DATA_BLOCK "DB_Z201_HMI"   // DB2010
{ S7_Optimized_Access := 'FALSE' }
VERSION : 0.1
   VAR
      tAlm : Struct   // HMI Alarms
         tE : Struct   // Emergency alarms
            xMainEmergency : Bool := TRUE;   // A122KE1.Main emergency ON {X|X|X|X|O}
            xSpare_1 : Bool := TRUE;
            xSpare_2 : Bool := TRUE;
            xSpare_3 : Bool := TRUE;
            xSpare_4 : Bool := TRUE;
            xSpare_5 : Bool := TRUE;
            xLocalMain1 : Bool := TRUE;   // A118SB1.Emergency localization MCC1201 {X|X|X|X|O}
            xLocalMain2 : Bool := TRUE;   // A118SB2.Emergency localization CS4201 {X|X|X|X|O}
            xLocalMain3 : Bool := TRUE;   // M204SSB3.Emergency localization M204S {X|X|X|X|O}
            xLocalMain4 : Bool := TRUE;   // M204SSB4.Emergency localization M204S {X|X|X|X|O}
            xLocalMain5 : Bool := FALSE;   // M211SB1.Emergency localization M211 {X|X|X|X|O}
            xLocalMain6 : Bool := FALSE;   // M211SB2.Emergency localization M211 {X|X|X|X|O}
            xLocalMain7 : Bool := FALSE;   // M218SB1.Emergency localization M218 {X|X|X|X|O}
            xLocalMain8 : Bool := FALSE;   // M218SB2.Emergency localization M218 {X|X|X|X|O}
            xLocalMain9 : Bool := FALSE;   // M214SB1.Emergency localization M214 {X|X|X|X|O}
            xLocalMain10 : Bool := FALSE;   // M214SB2.Emergency localization M214 {X|X|X|X|O}
            xLocalMain11 : Bool := FALSE;   // M203SB1.Emergency localization M203 {X|X|X|X|O}
            xLocalMain12 : Bool := FALSE;   // AxxSBx.Emergency localization Spare {X|X|X|X|O}
            xLocalMain13 : Bool := FALSE;   // AxxSBx.Emergency localization Spare {X|X|X|X|O}
            xSpare_19 : Bool := FALSE;
            xEmergencyONArea201 : Bool := FALSE;   // Emergency ON Area 201
            xEmergencyONArea301 : Bool := FALSE;   // Emergency ON Area 301
            xEmergencyONArea302 : Bool := FALSE;   // Emergency ON Area 302
            xEmergencyONArea501 : Bool := FALSE;   // Emergency ON Area 501
            xEmergencyONArea601 : Bool := FALSE;   // Emergency ON Area 601
            xEmergencyONArea701 : Bool := FALSE;   // Emergency ON Area 701
            xEmergencyONArea303 : Bool := FALSE;   // Emergency ON Area 303
            xSpare_27 : Bool := FALSE;
            xSpare_28 : Bool := FALSE;
            xSpare_29 : Bool := FALSE;
            xSpare_30 : Bool := FALSE;
            xSpare_31 : Bool := FALSE;
         END_STRUCT;
         tS : Struct   // Stopping faults
            xZ300NotReady : Bool := FALSE;   // Area 300 is not ready {X|X|X|X|O}
            xSpare_1 : Bool := FALSE;
            xSpare_2 : Bool := FALSE;
            xSpare_3 : Bool := FALSE;
            xSpare_4 : Bool := FALSE;
            xSpare_5 : Bool := FALSE;
            xSpare_6 : Bool := FALSE;
            xSpare_7 : Bool := FALSE;
            xSpare_8 : Bool := FALSE;
            xSpare_9 : Bool := FALSE;
            xSpare_10 : Bool := FALSE;
            xSpare_11 : Bool := FALSE;
            xSpare_12 : Bool := FALSE;
            xSpare_13 : Bool := FALSE;
            xSpare_14 : Bool := FALSE;
            xSpare_15 : Bool := FALSE;
            xSpare_16 : Bool := FALSE;
            xSpare_17 : Bool := FALSE;
            xSpare_18 : Bool := FALSE;
            xSpare_19 : Bool := FALSE;
            xSpare_20 : Bool := FALSE;
            xSpare_21 : Bool := FALSE;
            xSpare_22 : Bool := FALSE;
            xSpare_23 : Bool := FALSE;
            xSpare_24 : Bool := FALSE;
            xSpare_25 : Bool := FALSE;
            xSpare_26 : Bool := FALSE;
            xSpare_27 : Bool := FALSE;
            xSpare_28 : Bool := FALSE;
            xSpare_29 : Bool := FALSE;
            xSpare_30 : Bool := FALSE;
            xSpare_31 : Bool := FALSE;
         END_STRUCT;
         tF : Struct   // Faults
            xPowerFailure230vAux : Bool := FALSE;   // NU_A10QF1/2.Power failure 230v auxiliary / R13QF1.R13QF2.Power failure 230v auxiliary
            xPowerSupply24vLogic : Bool := FALSE;   // A109QF2.Power supply 24v logic / R18QF3.Power supply 24v logic
            xPowerSupply24vLogic2 : Bool := FALSE;   // A109QF3.Power supply 24v logic / R18QF4.Power supply 24v logic
            xPowerSuppluyOut24vUnderUpsEmOk : Bool := FALSE;   // A108QF5.Out24vUnderUpsEmOk / R18AP1.Redundancy 24v ok
            xPowerSupply24vLogic3 : Bool := FALSE;   // NU_A19QF1.Power supply 24v logic
            xPowerSupply24vLogic4 : Bool := FALSE;   // NU_A19QF2.Power supply 24v logic
            xPowerSuppluyOut24vUnderEmOk : Bool := FALSE;   // A108QF6.Out24vUnderEmOk
            xSpare_7 : Bool := FALSE;
            xPowerSupply24vDrive2 : Bool := FALSE;   // NU_A20QF4.Power Supply 24V Drive
            xSpare_9 : Bool := FALSE;
            xDriveSupply2 : Bool := FALSE;   // A137QM1.Drive Supply
            xSpare_11 : Bool := FALSE;
            xM216FanProtection : Bool;   // M216.A141QM1.Fan protection
            xM216FanFeedback : Bool;   // M216.A141KM1.Feedback rotation / M250.R12KM1.Feedback rotation
            xM209FanFeedback : Bool;   // M209.A178KM1.Feedback Rotation
            xSpare_15 : Bool;
            xSpare_16 : Bool;
            xSpare_17 : Bool;   // R204SP1.Compressed air presence cutting bridges
            xSpare_18 : Bool;
            xSpare_19 : Bool;
            xSpare_20 : Bool := FALSE;
            xSpare_21 : Bool := FALSE;
            xSpare_22 : Bool := FALSE;
            xSpare_23 : Bool := FALSE;
            xSpare_24 : Bool := FALSE;
            xSpare_25 : Bool := FALSE;
            xSpare_26 : Bool := FALSE;
            xSpare_27 : Bool := FALSE;
            xSpare_28 : Bool := FALSE;
            xSpare_29 : Bool := FALSE;
            xSpare_30 : Bool := FALSE;
            xSpare_31 : Bool := FALSE;
         END_STRUCT;
         tW : Struct   // Warnings
            xSpare_0 : Bool := FALSE;
            xSpare_1 : Bool := FALSE;
            xSpare_2 : Bool := FALSE;
            xSpare_3 : Bool := FALSE;
            xSpare_4 : Bool := FALSE;
            xSpare_5 : Bool := FALSE;
            xSpare_6 : Bool := FALSE;
            xSpare_7 : Bool := FALSE;
            xSpare_8 : Bool := FALSE;
            xSpare_9 : Bool := FALSE;
            xSpare_10 : Bool := FALSE;
            xSpare_11 : Bool := FALSE;
            xSpare_12 : Bool := FALSE;
            xSpare_13 : Bool := FALSE;
            xSpare_14 : Bool := FALSE;
            xSpare_15 : Bool := FALSE;
            xSpare_16 : Bool := FALSE;
            xSpare_17 : Bool := FALSE;
            xSpare_18 : Bool := FALSE;
            xSpare_19 : Bool := FALSE;
            xSpare_20 : Bool := FALSE;
            xSpare_21 : Bool := FALSE;
            xSpare_22 : Bool := FALSE;
            xSpare_23 : Bool := FALSE;
            xSpare_24 : Bool := FALSE;
            xSpare_25 : Bool := FALSE;
            xSpare_26 : Bool := FALSE;
            xSpare_27 : Bool := FALSE;
            xSpare_28 : Bool := FALSE;
            xSpare_29 : Bool := FALSE;
            xSpare_30 : Bool := FALSE;
            xSpare_31 : Bool := FALSE;
         END_STRUCT;
      END_STRUCT;
      tHMR : Struct   // HMI Read
         xSpare0 : Bool;
         xSpare1 : Bool;
         xSpare2 : Bool;
         xSpare3 : Bool;
         xSpare4 : Bool;
         xSpare5 : Bool;
         xSpare6 : Bool;
         xSpare7 : Bool;
         xSpare8 : Bool;
         xSpare9 : Bool;
         xSpare10 : Bool;
         xSpare11 : Bool;
         xSpare12 : Bool;
         xSpare13 : Bool;
         xSpare14 : Bool;
         xZoneAlarm : Bool := FALSE;   // Zone alarm {X|X|X|X|O}
         xSpare16 : Bool;
         xSpare17 : Bool;
         xSpare18 : Bool;
         xSpare19 : Bool;
         xSpare20 : Bool;
         xSpare21 : Bool;
         xSpare22 : Bool;
         xSpare23 : Bool;
         xSpare24 : Bool;
         xSpare25 : Bool;
         xSpare26 : Bool;
         xSpare27 : Bool;
         xSpare28 : Bool;
         xSpare29 : Bool;
         xSpare30 : Bool;
         xSpare31 : Bool;
         xSpare : Array[0..15] of Bool;
         iSpare0 : Int;
         iSpare1 : Int;
         iSpare2 : Int;
         iSpare3 : Int;
         iSpare4 : Int;
         iSpare5 : Int;
         iSpare6 : Int;
         iSpare7 : Int;
         iSpare8 : Int;
         iSpare9 : Int;
         iSpare10 : Int;
         iSpare11 : Int;
         iSpare12 : Int;
         iSpare13 : Int;
         iSpare14 : Int;
         iSpare15 : Int;
         iSpare16 : Int;
         dSpare0 : DInt;
         dZoneState : DInt := 1024;   // Zone status (1=CycleON 2=StopCyc 4=CycleReq 8=StopReq 1024=E-Stop) {X|X|X|X|O} / HMI Alarms
         dCabinetStatusMCC : DInt := 1;   // Cabinet status MCC1201 (1=OK;2=General power alarm;3=Local power alarm) {X|X|X|X|O} / HMI Write
         dDistanceFromSnaproll_cmm_M209 : DInt;   // Distance from snaproll [mm/100] {mm/100|mm|0|60000|M}
         dDistanceFromSnaproll_cmm_M216 : DInt;   // Distance from snaproll [mm/100] {mm/100|mm|0|60000|M}
         dSpare5 : DInt;
         dSpare6 : DInt;
         dSpare7 : DInt;
         dSpare8 : DInt;
         dSpare9 : DInt;
         dSpare10 : DInt;
         dSpare11 : DInt;
         dSpare12 : DInt;
         dSpare13 : DInt;
         dSpare14 : DInt;
         dSpare15 : DInt;
         rSpare0 : Real;
         rSpare1 : Real;
         rSpare2 : Real;
         rSpare3 : Real;
         rSpare4 : Real;
         rSpare5 : Real;
         rSpare6 : Real;
         rSpare7 : Real;
         rSpare8 : Real;
         tManCmd : Struct
            xFdbkRunFw : Bool;   // Feedback rotation FW all conveyors {x|x|x|x|O}
            xSpare1 : Bool;
            xSpare2 : Bool;
            xSpare3 : Bool;
            xSpare4 : Bool;
            xSpare5 : Bool;
            xSpare6 : Bool;
            xSpare7 : Bool;
            xSpare8 : Bool;
            xSpare9 : Bool;
            xSpare10 : Bool;
            xSpare11 : Bool;
            xSpare12 : Bool;
            xSpare13 : Bool;
            xSpare14 : Bool;
            xSpare15 : Bool;
            xSpare : Array[0..15] of Bool;
         END_STRUCT;
      END_STRUCT;
      tHMW : Struct   // HMI Write
         xSpare0 : Bool;
         xSpare1 : Bool;
         xSpare2 : Bool;
         xSpare3 : Bool;
         xSpare4 : Bool;
         xStartCycleRequest : Bool := FALSE;   // Start cycle request {X|X|X|X|O}
         xStopCycleRequest : Bool := FALSE;   // Stop cycle request {X|X|X|X|O}
         xForceStopCycle : Bool := FALSE;   // Force stop cycle {X|X|X|X|O}
         xSpare8 : Bool;
         xEnabledChipsBlowerM216 : Bool;   // Chips Blower M216 Enabled {X|X|X|X|O}
         xEnabledChipsBlowerM209 : Bool;   // Chips Blower M209 Enabled {X|X|X|X|O}
         xUpdateDistSnap_M209 : Bool;   // Update distance from snap roll {x|x|x|x|M}
         xUpdateDistSnap_M216 : Bool;
         xSpare13 : Bool;
         xEnableManualCommand : Bool;   // Enable Disable Manual command {x|x|x|x|O}
         xFaultsReset : Bool := FALSE;   // Reset faults {X|X|X|X|O}
         xGeneralReset : Bool := FALSE;   // General reset {X|X|X|X|M}
         xSpare17 : Bool;
         xSpare18 : Bool;
         xSpare19 : Bool;
         xSpare20 : Bool;
         xSpare21 : Bool;
         xSpare22 : Bool;
         xSpare23 : Bool;
         xSpare24 : Bool;
         xSpare25 : Bool;
         xSpare26 : Bool;
         xSpare27 : Bool;
         xSpare28 : Bool;
         xSpare29 : Bool;
         xSpare30 : Bool;
         xSpare31 : Bool;
         xSpare : Array[0..15] of Bool;
         iSpare0 : Int;
         iSpare1 : Int;
         iSpare2 : Int;
         iSpare3 : Int;
         iSpare4 : Int;
         iSpare5 : Int;
         iSpare6 : Int;
         iSpare7 : Int;
         iSpare8 : Int;
         iSpare9 : Int;
         iSpare10 : Int;
         iSpare11 : Int;
         iSpare12 : Int;
         iSpare13 : Int;
         iSpare14 : Int;
         iSpare15 : Int;
         iSpare16 : Int;
         dDistanceFromSnaproll_cmm_M209 : DInt;   // Distance from snaproll [mm/100] [mm/100] {mm/100|mm|0|60000|M}
         dDistanceFromSnaproll_cmm_M216 : DInt;   // Distance from snaproll [mm/100] [mm/100] {mm/100|mm|0|60000|M}
         dSpare2 : DInt;
         dSpare3 : DInt;
         dSpare4 : DInt;
         dSpare5 : DInt;
         dSpare6 : DInt;
         dSpare7 : DInt;
         dSpare8 : DInt;
         dSpare9 : DInt;
         dSpare10 : DInt;
         dSpare11 : DInt;
         dSpare12 : DInt;
         dSpare13 : DInt;
         dSpare14 : DInt;
         dSpare15 : DInt;
         dSpare16 : DInt;
         rSpare0 : Real;
         rSpare1 : Real;
         rSpare2 : Real;
         rSpare3 : Real;
         rSpare4 : Real;
         rSpare5 : Real;
         rSpare6 : Real;
         rSpare7 : Real;
         rSpare8 : Real;
         tManCmd : Struct
            xRunFw : Bool;   // Rotation FW all conveyors {x|x|x|x|O}
            xSpare1 : Bool;
            xSpare2 : Bool;
            xSpare3 : Bool;
            xSpare4 : Bool;
            xSpare5 : Bool;
            xSpare6 : Bool;
            xSpare7 : Bool;
            xSpare8 : Bool;
            xSpare9 : Bool;
            xSpare10 : Bool;
            xSpare11 : Bool;
            xSpare12 : Bool;
            xSpare13 : Bool;
            xSpare14 : Bool;
            xSpare15 : Bool;
            xSpare16 : Bool;
            xSpare17 : Bool;
            xSpare18 : Bool;
            xSpare19 : Bool;
            xSpare20 : Bool;
            xSpare21 : Bool;
            xSpare22 : Bool;
            xSpare23 : Bool;
            xSpare24 : Bool;
            xSpare25 : Bool;
            xSpare26 : Bool;
            xSpare27 : Bool;
            xSpare28 : Bool;
            xSpare29 : Bool;
            xSpare30 : Bool;
            xSpare31 : Bool;
         END_STRUCT;
      END_STRUCT;
   END_VAR
BEGIN
END_DATA_BLOCK

DATA_BLOCK "DB_ZUPS_HMI"   // DB2012
{ S7_Optimized_Access := 'FALSE' }
VERSION : 0.1
   VAR
      tAlm : Struct   // HMI Alarms
         tE : Struct   // Emergency alarms
            xSpare_0 : Bool := TRUE;
            xMainEmergencyUPS : Bool := TRUE;   // A117KE1.Main emergency UPS ON {X|X|X|X|O}
            xLocalUPS1 : Bool := TRUE;   // AxxSB1.Emergency localization MCC1201 {X|X|X|X|O}
            xLocalUPS2 : Bool := TRUE;   // M204S_SB1.Emergency localization M204S {X|X|X|X|O}
            xLocalUPS3 : Bool := TRUE;   // M204S_SB2.Emergency localization M204S {X|X|X|X|O}
            xLocalUPS4 : Bool := TRUE;   // CS4201A117SB1.Emergency localization spare {X|X|X|X|O}
            xLocalUpS5 : Bool := TRUE;   // AxxSBx.Emergency localization spare {X|X|X|X|O}
            xSpare_7 : Bool := TRUE;
            xSpare_8 : Bool := TRUE;
            xSpare_9 : Bool := TRUE;
            xSpare_10 : Bool := FALSE;
            xSpare_11 : Bool := FALSE;
            xSpare_12 : Bool := FALSE;
            xSpare_13 : Bool := FALSE;
            xSpare_14 : Bool := FALSE;
            xSpare_15 : Bool := FALSE;
            xSpare_16 : Bool := FALSE;
            xSpare_17 : Bool := FALSE;
            xSpare_18 : Bool := FALSE;
            xSpare_19 : Bool := FALSE;
            xSpare_20 : Bool := FALSE;
            xSpare_21 : Bool := FALSE;
            xSpare_22 : Bool := FALSE;
            xSpare_23 : Bool := FALSE;
            xSpare_24 : Bool := FALSE;
            xSpare_25 : Bool := FALSE;
            xSpare_26 : Bool := FALSE;
            xSpare_27 : Bool := FALSE;
            xSpare_28 : Bool := FALSE;
            xSpare_29 : Bool := FALSE;
            xSpare_30 : Bool := FALSE;
            xSpare_31 : Bool := FALSE;
         END_STRUCT;
         tS : Struct   // Stopping faults
            xSpare_0 : Bool := FALSE;
            xSpare_1 : Bool := FALSE;
            xSpare_2 : Bool := FALSE;
            xSpare_3 : Bool := FALSE;
            xSpare_4 : Bool := FALSE;
            xSpare_5 : Bool := FALSE;
            xSpare_6 : Bool := FALSE;
            xSpare_7 : Bool := FALSE;
            xSpare_8 : Bool := FALSE;
            xSpare_9 : Bool := FALSE;
            xSpare_10 : Bool := FALSE;
            xSpare_11 : Bool := FALSE;
            xSpare_12 : Bool := FALSE;
            xSpare_13 : Bool := FALSE;
            xSpare_14 : Bool := FALSE;
            xSpare_15 : Bool := FALSE;
            xSpare_16 : Bool := FALSE;
            xSpare_17 : Bool := FALSE;
            xSpare_18 : Bool := FALSE;
            xSpare_19 : Bool := FALSE;
            xSpare_20 : Bool := FALSE;
            xSpare_21 : Bool := FALSE;
            xSpare_22 : Bool := FALSE;
            xSpare_23 : Bool := FALSE;
            xSpare_24 : Bool := FALSE;
            xSpare_25 : Bool := FALSE;
            xSpare_26 : Bool := FALSE;
            xSpare_27 : Bool := FALSE;
            xSpare_28 : Bool := FALSE;
            xSpare_29 : Bool := FALSE;
            xSpare_30 : Bool := FALSE;
            xSpare_31 : Bool := FALSE;
         END_STRUCT;
         tF : Struct   // Faults
            xSpare_0 : Bool := FALSE;   // R13QF1.R13QF2.Power failure 230v auxiliary
            xSpare_1 : Bool := FALSE;   // R18QF3.Power supply 24v logic
            xSpare_2 : Bool := FALSE;   // R18QF4.Power supply 24v logic
            xSpare_3 : Bool := FALSE;   // R18AP1.Redundancy 24v ok
            xSpare_4 : Bool := FALSE;
            xSpare_5 : Bool := FALSE;
            xSpare_6 : Bool := FALSE;
            xPowerSupply24vDrive1 : Bool := FALSE;   // A110QF2.Power Supply 24V Drive
            xSpare_8 : Bool := FALSE;
            xDriveSupply1 : Bool := FALSE;   // A136QM1.Drive Supply
            xSpare_10 : Bool := FALSE;
            xSpare_11 : Bool := FALSE;
            xSpare_12 : Bool;
            xSpare_13 : Bool;   // M250.R12KM1.Feedback rotation
            xSpare_14 : Bool;
            xSpare_15 : Bool;
            xSpare_16 : Bool;
            xSpare_17 : Bool;   // R204SP1.Compressed air presence cutting bridges
            xSpare_18 : Bool;
            xSpare_19 : Bool;
            xSpare_20 : Bool := FALSE;
            xSpare_21 : Bool := FALSE;
            xSpare_22 : Bool := FALSE;
            xSpare_23 : Bool := FALSE;
            xSpare_24 : Bool := FALSE;
            xSpare_25 : Bool := FALSE;
            xSpare_26 : Bool := FALSE;
            xSpare_27 : Bool := FALSE;
            xSpare_28 : Bool := FALSE;
            xSpare_29 : Bool := FALSE;
            xSpare_30 : Bool := FALSE;
            xSpare_31 : Bool := FALSE;
         END_STRUCT;
         tW : Struct   // Warnings
            xSpare_0 : Bool := FALSE;
            xSpare_1 : Bool := FALSE;
            xSpare_2 : Bool := FALSE;
            xSpare_3 : Bool := FALSE;
            xSpare_4 : Bool := FALSE;
            xSpare_5 : Bool := FALSE;
            xSpare_6 : Bool := FALSE;
            xSpare_7 : Bool := FALSE;
            xSpare_8 : Bool := FALSE;
            xSpare_9 : Bool := FALSE;
            xSpare_10 : Bool := FALSE;
            xSpare_11 : Bool := FALSE;
            xSpare_12 : Bool := FALSE;
            xSpare_13 : Bool := FALSE;
            xSpare_14 : Bool := FALSE;
            xSpare_15 : Bool := FALSE;
            xSpare_16 : Bool := FALSE;
            xSpare_17 : Bool := FALSE;
            xSpare_18 : Bool := FALSE;
            xSpare_19 : Bool := FALSE;
            xSpare_20 : Bool := FALSE;
            xSpare_21 : Bool := FALSE;
            xSpare_22 : Bool := FALSE;
            xSpare_23 : Bool := FALSE;
            xSpare_24 : Bool := FALSE;
            xSpare_25 : Bool := FALSE;
            xSpare_26 : Bool := FALSE;
            xSpare_27 : Bool := FALSE;
            xSpare_28 : Bool := FALSE;
            xSpare_29 : Bool := FALSE;
            xSpare_30 : Bool := FALSE;
            xSpare_31 : Bool := FALSE;
         END_STRUCT;
      END_STRUCT;
      tHMR : Struct   // HMI Read
         xSpare0 : Bool;
         xSpare1 : Bool;
         xSpare2 : Bool;
         xSpare3 : Bool;
         xSpare4 : Bool;
         xSpare5 : Bool;
         xSpare6 : Bool;
         xSpare7 : Bool;
         xSpare8 : Bool;
         xSpare9 : Bool;
         xSpare10 : Bool;
         xSpare11 : Bool;
         xSpare12 : Bool;
         xSpare13 : Bool;
         xSpare14 : Bool;
         xZoneAlarm : Bool := FALSE;   // Zone alarm {X|X|X|X|O}
         xSpare16 : Bool;
         xSpare17 : Bool;
         xSpare18 : Bool;
         xSpare19 : Bool;
         xSpare20 : Bool;
         xSpare21 : Bool;
         xSpare22 : Bool;
         xSpare23 : Bool;
         xSpare24 : Bool;
         xSpare25 : Bool;
         xSpare26 : Bool;
         xSpare27 : Bool;
         xSpare28 : Bool;
         xSpare29 : Bool;
         xSpare30 : Bool;
         xSpare31 : Bool;
         xSpare : Array[0..15] of Bool;
         iSpare0 : Int;
         iSpare1 : Int;
         iSpare2 : Int;
         iSpare3 : Int;
         iSpare4 : Int;
         iSpare5 : Int;
         iSpare6 : Int;
         iSpare7 : Int;
         iSpare8 : Int;
         iSpare9 : Int;
         iSpare10 : Int;
         iSpare11 : Int;
         iSpare12 : Int;
         iSpare13 : Int;
         iSpare14 : Int;
         iSpare15 : Int;
         iSpare16 : Int;
         dSpare0 : DInt;
         dZoneState : DInt := 1024;   // Zone status (1=CycleON 2=StopCyc 4=CycleReq 8=StopReq 1024=E-Stop) {X|X|X|X|O} / HMI Alarms
         dSpare2 : DInt;
         dSpare3 : DInt;
         dSpare4 : DInt;
         dSpare5 : DInt;
         dSpare6 : DInt;
         dSpare7 : DInt;
         dSpare8 : DInt;
         dSpare9 : DInt;
         dSpare10 : DInt;
         dSpare11 : DInt;
         dSpare12 : DInt;
         dSpare13 : DInt;
         dSpare14 : DInt;
         dSpare15 : DInt;
         rSpare0 : Real;
         rSpare1 : Real;
         rSpare2 : Real;
         rSpare3 : Real;
         rSpare4 : Real;
         rSpare5 : Real;
         rSpare6 : Real;
         rSpare7 : Real;
         rSpare8 : Real;
         tManCmd : Struct
            xSpare0 : Bool;
            xSpare1 : Bool;
            xSpare2 : Bool;
            xSpare3 : Bool;
            xSpare4 : Bool;
            xSpare5 : Bool;
            xSpare6 : Bool;
            xSpare7 : Bool;
            xSpare8 : Bool;
            xSpare9 : Bool;
            xSpare10 : Bool;
            xSpare11 : Bool;
            xSpare12 : Bool;
            xSpare13 : Bool;
            xSpare14 : Bool;
            xSpare15 : Bool;
            xSpare : Array[0..15] of Bool;
         END_STRUCT;
      END_STRUCT;
      tHMW : Struct   // HMI Write
         xSpare0 : Bool;
         xSpare1 : Bool;
         xSpare2 : Bool;
         xSpare3 : Bool;
         xSpare4 : Bool;
         xStartCycleRequest : Bool := FALSE;   // Start cycle request {X|X|X|X|O}
         xStopCycleRequest : Bool := FALSE;   // Stop cycle request {X|X|X|X|O}
         xForceStopCycle : Bool := FALSE;   // Force stop cycle {X|X|X|X|O}
         xSpare8 : Bool;
         xSpare9 : Bool;
         xSpare10 : Bool;
         xSpare11 : Bool;
         xSpare12 : Bool;
         xSpare13 : Bool;
         xSpare14 : Bool;
         xFaultsReset : Bool := FALSE;   // Reset faults {X|X|X|X|O}
         xSpare16 : Bool := FALSE;
         xSpare17 : Bool;
         xSpare18 : Bool;
         xSpare19 : Bool;
         xSpare20 : Bool;
         xSpare21 : Bool;
         xSpare22 : Bool;
         xSpare23 : Bool;
         xSpare24 : Bool;
         xSpare25 : Bool;
         xSpare26 : Bool;
         xSpare27 : Bool;
         xSpare28 : Bool;
         xSpare29 : Bool;
         xSpare30 : Bool;
         xSpare31 : Bool;
         xSpare : Array[0..15] of Bool;
         iSpare0 : Int;
         iSpare1 : Int;
         iSpare2 : Int;
         iSpare3 : Int;
         iSpare4 : Int;
         iSpare5 : Int;
         iSpare6 : Int;
         iSpare7 : Int;
         iSpare8 : Int;
         iSpare9 : Int;
         iSpare10 : Int;
         iSpare11 : Int;
         iSpare12 : Int;
         iSpare13 : Int;
         iSpare14 : Int;
         iSpare15 : Int;
         iSpare16 : Int;
         dSpare0 : DInt;
         dSpare1 : DInt;
         dSpare2 : DInt;
         dSpare3 : DInt;
         dSpare4 : DInt;
         dSpare5 : DInt;
         dSpare6 : DInt;
         dSpare7 : DInt;
         dSpare8 : DInt;
         dSpare9 : DInt;
         dSpare10 : DInt;
         dSpare11 : DInt;
         dSpare12 : DInt;
         dSpare13 : DInt;
         dSpare14 : DInt;
         dSpare15 : DInt;
         dSpare16 : DInt;
         rSpare0 : Real;
         rSpare1 : Real;
         rSpare2 : Real;
         rSpare3 : Real;
         rSpare4 : Real;
         rSpare5 : Real;
         rSpare6 : Real;
         rSpare7 : Real;
         rSpare8 : Real;
         tManCmd : Struct
            xSpare0 : Bool;
            xSpare1 : Bool;
            xSpare2 : Bool;
            xSpare3 : Bool;
            xSpare4 : Bool;
            xSpare5 : Bool;
            xSpare6 : Bool;
            xSpare7 : Bool;
            xSpare8 : Bool;
            xSpare9 : Bool;
            xSpare10 : Bool;
            xSpare11 : Bool;
            xSpare12 : Bool;
            xSpare13 : Bool;
            xSpare14 : Bool;
            xSpare15 : Bool;
            xSpare16 : Bool;
            xSpare17 : Bool;
            xSpare18 : Bool;
            xSpare19 : Bool;
            xSpare20 : Bool;
            xSpare21 : Bool;
            xSpare22 : Bool;
            xSpare23 : Bool;
            xSpare24 : Bool;
            xSpare25 : Bool;
            xSpare26 : Bool;
            xSpare27 : Bool;
            xSpare28 : Bool;
            xSpare29 : Bool;
            xSpare30 : Bool;
            xSpare31 : Bool;
         END_STRUCT;
      END_STRUCT;
   END_VAR
BEGIN
END_DATA_BLOCK

// folder: TaskMedium

DATA_BLOCK "FB_OptManager_V1_00_IDB"   // DB7
{ S7_Optimized_Access := 'TRUE' }
VERSION : 0.1
// stored: InstanceOfName FB_OptManager_V1.00
"FB_OptManager_V1.00"
BEGIN
END_DATA_BLOCK

DATA_BLOCK "GP_OB_Initialize_Medium_IDB"   // DB9
{ S7_Optimized_Access := 'TRUE' }
AUTHOR : Cigliutt
FAMILY : GP
VERSION : 1.1
// stored: InstanceOfName GP_OB_Initialize
"GP_OB_Initialize"
BEGIN
END_DATA_BLOCK

DATA_BLOCK "GP_OB_Initialize_Slow_IDB"   // DB10
{ S7_Optimized_Access := 'TRUE' }
AUTHOR : Cigliutt
FAMILY : GP
VERSION : 1.1
// stored: InstanceOfName GP_OB_Initialize
"GP_OB_Initialize"
BEGIN
END_DATA_BLOCK

DATA_BLOCK "FB_Snaproll_V1_00_IDB"   // DB21
{ S7_Optimized_Access := 'TRUE' }
VERSION : 0.1
// stored: InstanceOfName FB_Snaproll_V1.00
"FB_Snaproll_V1.00"
BEGIN
END_DATA_BLOCK

DATA_BLOCK "FB_CommunicationZ300_V1.00_DB_1"   // DB25
{ S7_Optimized_Access := 'TRUE' }
VERSION : 0.1
// stored: InstanceOfName FB_CommunicationZ300_V1.00
"FB_CommunicationZ300_V1.00"
BEGIN
END_DATA_BLOCK

DATA_BLOCK "FB_CommunicationZ300_V1.00_DB"   // DB28
{ S7_Optimized_Access := 'TRUE' }
VERSION : 0.1
// stored: InstanceOfName FB_CommunicationZ300_V1.00
"FB_CommunicationZ300_V1.00"
BEGIN
END_DATA_BLOCK

DATA_BLOCK "FB_Defects_Add_Medium_V1_00_IDB"   // DB36
{ S7_Optimized_Access := 'TRUE' }
VERSION : 0.1
// stored: InstanceOfName FB_Defects_Add_V1.00
"FB_Defects_Add_V1.00"
BEGIN
END_DATA_BLOCK

// folder: TaskSlow

DATA_BLOCK "FB_Digitizer_2_V1_00_IDB"   // DB11
{ S7_Optimized_Access := 'TRUE' }
VERSION : 0.1
// stored: InstanceOfName FB_Digitizer_V1.00
"FB_Digitizer_V1.00"
BEGIN
END_DATA_BLOCK

DATA_BLOCK "FB_Digitizer_1_V1_00_IDB"   // DB12
{ S7_Optimized_Access := 'TRUE' }
VERSION : 0.1
// stored: InstanceOfName FB_Digitizer_V1.00
"FB_Digitizer_V1.00"
BEGIN
END_DATA_BLOCK

DATA_BLOCK "Z200"   // DB13
{ S7_Optimized_Access := 'TRUE' }
VERSION : 0.1
   VAR
      tmON_24Vdc : "UDT_IECTON_V1.00";   // Presence 24Vdc timer / 24VDC ok delayed timer
      ST_xZoneError : Bool := FALSE;   // Zone error / Zone is in error
      ST_xFaultsEnabled : Bool := TRUE;   // Faults enabled
      ST_xZoneFaults : Bool := TRUE;   // Cumulative of zone faults / Zone is in faults
      ST_xZoneStoppingFaults : Bool := FALSE;   // Cumulative of zone stopping faults / Zone is in stopping faults
      ST_xOutputEnabledM250Fan : Bool;   // Output enable M250 fan
      ST_xOutputEnabledM272Chips : Bool;   // Output enable M272 chips blower
      ST_xOutputEnabledM220Brush : Bool;   // Output enable M272 chips blower
      ST_xZoneWarnings : Bool := FALSE;   // Cumulative of zone warning / Zone is in warning
      ST_xCycleON : Bool := TRUE;   // Zone in cycle ON / Cycle ON
      ST_xConditionOKStopCycle : Bool := TRUE;   // Condition ok to accept stop cycle
      ST_xCycleONDelayed : Bool := TRUE;   // Cycle ON delayed
      ST_xConditionOkPhaseAdvancement : Bool := FALSE;   // Condition ok for phase advancement
      ST_xConditionOkCycleON : Bool := FALSE;   // Condition ok for cycle ON
      ST_xMachineReset : Bool := FALSE;   // Machine reset request
      ST_xPLC1 : Bool := TRUE;   // This is PLC 1
      ST_xPLC2 : Bool := FALSE;   // This is PLC 2
      ST_xThisPlcActive : Bool := TRUE;   // This PLC is active
      ST_xStartCycleRequest : Bool := FALSE;   // Request start cycle
      ST_xStopCycleRequest : Bool := FALSE;   // Request stop cycle
      ST_xM209GlassBreak : Bool;   // M272 Chips blower glass break
      ST_xM203GlassBreak : Bool;   // M272 Chips blower glass break
      OSR_xStartCycle : Bool := FALSE;   // OSR start cycle
      OSR_xStopCycle : Bool := FALSE;   // OSR stop cycle
      OSR_xForceStopCycle : Bool := FALSE;   // OSR force stop cycle
      OSR_xChipsBlowerON : Bool;   // OSR chips blower on
      OSR_xSBResetAnomaly : Bool;   // OSR reset anomaly
      OS_xStartCycle : Bool := FALSE;   // OS start cycle
      OS_xStopCycle : Bool := FALSE;   // OS stop cycle
      OS_xForceStopCycle : Bool := FALSE;   // OS force stop cycle
      OS_xChipsBlowerON : Bool;   // OS chips blower on
      OS_xCpuActive : Bool;   // OS Cpu active
      OSR_xCpuActive : Bool;   // OSR Cpu active
      ST_xStopCycleAccepted : Bool := FALSE;   // Stop cycle accepted
      AUX_tmON_M250FanFeedback : "UDT_IECTON_V1.00";   // M250 Fan feedback anomaly
      tOutputs : Struct
         xPLC1On : Bool;   // o.A195AP1.A255HL4.EnableCPUA
         xPLC2On : Bool;   // o.A195AP1.A255HL5.EnableCPUB
         xEmergencyON : Bool;   // o.A195AP1.A255HL1/1A.EmergencyON
         xSafetiesON : Bool;   // o.A195AP1.A255HL3.SafetiesON
         xHLResetAnomaly : Bool;   // o.A195AP1.A207SB1.HLResetAnomalyZ200
         xHAAlarm : Bool;   // o.A401AP1.A416HA1.Alarm
      END_STRUCT;
      tInputs : Struct
         xPowerSupply230vAux : Bool := FALSE;   // i.A195AP1.A10QF1/2.PowerFailure230VAuxiliary / i.R195AP1.R13QF1/2.PowerFailure230VAuxiliary
         xRedundancy24vOk1 : Bool;   // i.R195AP1.R18AP1.Redundacy24VOk / i.A195AP1.A18AP1.Redundancy24VOk
         xPowerSupply24vProt1 : Bool;
         xPowerSupply24vProt2 : Bool;
         xProtectionCommandsAnomalies : Bool := FALSE;   // i.A195AP1.A18QF3.PowerSupply24VLogic / i.R195AP1.R18QF3.PowerSupply24VLogic
         xProtectionCommandsInternalInput : Bool := FALSE;   // i.A195AP1.A18QF4.PowerSupply24VLogic / i.R195AP1.R18QF4.PowerSupply24VLogic
         xProtectionCommandsInternalOutput : Bool := FALSE;   // i.A195AP1.A19QF1.PowerSupply24VLogic / i.R195AP1.R18QF4.PowerSupply24VLogic
         xProtectionCommandsExternalInput : Bool := FALSE;   // i.A195AP1.A19QF2.PowerSupply24VLogic / i.R195AP1.R18QF4.PowerSupply24VLogic
         xMainEmergencyON : Bool := FALSE;   // i.A195AP1.A45KE1.MainEmergencyON / i.R195AP1.R18QF4.PowerSupply24VLogic
         xCPUAEnabled : Bool := FALSE;   // i.A151AP1.Selection CPU A / i.R150AP1.CPU A Enabled
         xCPUBEnabled : Bool := TRUE;   // i.A151AP1.Selection CPU B / i.R150AP1.CPU B Enabled
         xCPUARecognition : Bool := FALSE;   // i.A151AP1.Recognition CPU A / i.R150AP1.Recognition CPU A
         xCPUBRecognition : Bool := FALSE;   // i.A151AP1.Recognition CPU B / i.R150AP1.Recognition CPU B
         xFeedbackSwitch : Bool;
         xFeedbackAbilitationCPU_B : Bool;
         xCompressedAirPresence : Bool;
         xSBResetAnomalyZ200 : Bool;   // i.A195AP1.A207SB1.ResetAnomalyZ200
      END_STRUCT;
   END_VAR
BEGIN
END_DATA_BLOCK

DATA_BLOCK "FB_DigitizerManager_V1_00_IDB"   // DB15
{ S7_Optimized_Access := 'TRUE' }
VERSION : 0.1
// stored: InstanceOfName FB_DigitizerManager_V1.00
"FB_DigitizerManager_V1.00"
BEGIN
END_DATA_BLOCK

DATA_BLOCK "FB_YCuts2_V1_00_IDB"   // DB16
{ S7_Optimized_Access := 'TRUE' }
VERSION : 0.1
// stored: InstanceOfName FB_YCuts_V1.00
"FB_YCuts_V1.00"
BEGIN
END_DATA_BLOCK

DATA_BLOCK "FB_CrossCuts_2_V1_00_IDB"   // DB19
{ S7_Optimized_Access := 'TRUE' }
VERSION : 0.1
// stored: InstanceOfName FB_CrossCutsModbus_V1.00
"FB_CrossCutsModbus_V1.00"
BEGIN
   tHMW.dOperStartCutPos_cmm := -150000;
   tHMW.dOperEndCutPos_cmm := 150000;
   tHMW.dDescReactTime_ms := 200;
   tHMW.dRaiseReactTime_ms := 30;
   tHMW.dFireONReactTime_ms := 200;
   tHMW.dFireOFFReactTime_ms := 5;
   tHMW.dCutStartOffsetDelay_cmm := -11000;
   tHMW.dCutEndOffsetDelay_cmm := 1000;
   tHMW.dDistanceFromSnaproll_cmm := 445500;
   tHMW.dAngleValue_uDegree := 9500000;
   tHMW.dDistanceFromCenterLine_cmm := -290000;
   tHMW.dDistTeoLength_cmm := 200000;
   tHMW.dDistRealLength_cmm := 200050;
   tHMW.dCuttingPressure_mN := 20000;
   tHMW.dCutPriority := 2;
   tHMR.dActualCutPosRequest := 4;
   tHMR.dXCutStatusRequest := 3;
   tHMR.dXCutActualStatus := 3;
   tHMR.dDistanceFromSnaproll_cmm := 446100;
   tHMR.dAngleValue_uDegree := 9580000;
   tHMR.dDistanceFromCenterLine_cmm := -290000;
   tHMR.dStatus := 1;
   tHMR.rHeadUsage_km := 3.41702;
END_DATA_BLOCK

DATA_BLOCK "FB_CrossCuts_1_V1_00_IDB"   // DB20
{ S7_Optimized_Access := 'TRUE' }
VERSION : 0.1
// stored: InstanceOfName FB_CrossCutsModbus_V1.00
"FB_CrossCutsModbus_V1.00"
BEGIN
   tHMW.dOperStartCutPos_cmm := -180000;
   tHMW.dOperEndCutPos_cmm := 140000;
   tHMW.dDescReactTime_ms := 200;
   tHMW.dRaiseReactTime_ms := 30;
   tHMW.dFireONReactTime_ms := 200;
   tHMW.dFireOFFReactTime_ms := 5;
   tHMW.dCutStartOffsetDelay_cmm := -8000;
   tHMW.dCutEndOffsetDelay_cmm := 1000;
   tHMW.dDistanceFromSnaproll_cmm := 528000;
   tHMW.dAngleValue_uDegree := 9500000;
   tHMW.dDistanceFromCenterLine_cmm := -290000;
   tHMW.dDiagRealLength_cmm := 510000;
   tHMW.dDiagRealWidth_cmm := 315000;
   tHMW.dDiagGlassFlow_cmm := 599900;
   tHMW.dDiagGlassOppFlow_cmm := 598900;
   tHMW.dCuttingPressure_mN := 19000;
   tHMW.dCutPriority := 2;
   tHMR.dActualCutPosRequest := 4;
   tHMR.dXCutStatusRequest := 3;
   tHMR.dXCutActualStatus := 3;
   tHMR.dDistanceFromSnaproll_cmm := 528000;
   tHMR.dAngleValue_uDegree := 9600000;
   tHMR.dDistanceFromCenterLine_cmm := -290000;
   tHMR.dStatus := 1;
   tHMR.rHeadUsage_km := 45.7704;
END_DATA_BLOCK

DATA_BLOCK "FB_YCuts1_V1_00_IDB"   // DB22
{ S7_Optimized_Access := 'TRUE' }
VERSION : 0.1
// stored: InstanceOfName FB_YCuts_V1.00
"FB_YCuts_V1.00"
BEGIN
END_DATA_BLOCK

DATA_BLOCK "FB_Markers_V1.00_IDB"   // DB24
{ S7_Optimized_Access := 'TRUE' }
VERSION : 0.1
// stored: InstanceOfName FB_Markers_V1.00
"FB_Markers_V1.00"
BEGIN
END_DATA_BLOCK

DATA_BLOCK "FB_WanderCamera_V1_00_IDB"   // DB26
{ S7_Optimized_Access := 'TRUE' }
VERSION : 0.1
// stored: InstanceOfName FB_WanderCamera_V1.00
"FB_WanderCamera_V1.00"
BEGIN
END_DATA_BLOCK

DATA_BLOCK "FB_LehrSpeed_IDB"   // DB27
{ S7_Optimized_Access := 'TRUE' }
VERSION : 0.1
// stored: InstanceOfName FB_LehrSpeed
"FB_LehrSpeed"
BEGIN
END_DATA_BLOCK

DATA_BLOCK "FB_CrossCuts_3_V1_00_IDB"   // DB30
{ S7_Optimized_Access := 'TRUE' }
VERSION : 0.1
// stored: InstanceOfName FB_CrossCutsModbus_V1.00
"FB_CrossCutsModbus_V1.00"
BEGIN
END_DATA_BLOCK

DATA_BLOCK "FB_ColdBackupManager_V1_00_DB"   // DB32
{ S7_Optimized_Access := 'TRUE' }
VERSION : 0.1
// stored: InstanceOfName FB_ColdBackupManager_V1.00
"FB_ColdBackupManager_V1.00"
BEGIN
END_DATA_BLOCK

DATA_BLOCK "FB_Defects_Add_Slow_V1_00_IDB"   // DB37
{ S7_Optimized_Access := 'TRUE' }
VERSION : 0.1
// stored: InstanceOfName FB_Defects_Add_V1.00
"FB_Defects_Add_V1.00"
BEGIN
END_DATA_BLOCK

DATA_BLOCK "DataTime_HMI"   // DB42
{ S7_Optimized_Access := 'TRUE' }
VERSION : 0.1
   VAR RETAIN
      DTL_DataTime : DTL;
   END_VAR
BEGIN
END_DATA_BLOCK

DATA_BLOCK "FB_BD_BreakPH_V1_00_IDB"   // DB45
{ S7_Optimized_Access := 'TRUE' }
VERSION : 0.1
// stored: InstanceOfName FB_BreakDetector_V1.00
"FB_BreakDetector_V1.00"
BEGIN
END_DATA_BLOCK

DATA_BLOCK "FB_Oil_V1_00_IDB"   // DB49
{ S7_Optimized_Access := 'TRUE' }
VERSION : 0.1
// stored: InstanceOfName FB_Oil_V1.00
"FB_Oil_V1.00"
BEGIN
END_DATA_BLOCK

DATA_BLOCK "FB_ManInsp_V1_00_IDB"   // DB50
{ S7_Optimized_Access := 'TRUE' }
VERSION : 0.1
// stored: InstanceOfName FB_ManInsp_V1.00
"FB_ManInsp_V1.00"
BEGIN
END_DATA_BLOCK

DATA_BLOCK "FB_ISRA5D_IDB"   // DB55
{ S7_Optimized_Access := 'TRUE' }
VERSION : 0.1
// stored: InstanceOfName FB_ISRA5D
"FB_ISRA5D"
BEGIN
END_DATA_BLOCK

DATA_BLOCK "FB_CrossCut_Opt_V1_00_IDB"   // DB61
{ S7_Optimized_Access := 'TRUE' }
VERSION : 0.1
// stored: InstanceOfName FB_CrossCutOpt_V1.00
"FB_CrossCutOpt_V1.00"
BEGIN
END_DATA_BLOCK

DATA_BLOCK "FB_BD_DigitizerPH_V1_00_IDB"   // DB67
{ S7_Optimized_Access := 'TRUE' }
VERSION : 0.1
// stored: InstanceOfName FB_BreakDetector_V1.00
"FB_BreakDetector_V1.00"
BEGIN
END_DATA_BLOCK

// folder: 02_Inputs

FUNCTION "InputTaskFast" : Void   // FC8, LAD
{ S7_Optimized_Access := 'TRUE' }
VERSION : 0.1
BEGIN

REGION Network 2 (SCL)
   "FB_TrackEncoder_V1_00_IDB".INP_tHSCCount := "i_HSCInput_Count1";
END_REGION
END_FUNCTION

FUNCTION "InputTaskSlow" : Void   // FC9, LAD
{ S7_Optimized_Access := 'TRUE' }
VERSION : 0.1
   VAR_TEMP
      TMP_xToAssign : Bool;
   END_VAR
BEGIN

REGION Network 1 (SCL)
   //"ZUPS".tInputs.xEmergencyONAreaUPS := "i.A195AP1.A32KE1.EmergencyAreaUPSON";
   //"ZUPS".tInputs.xPowerSupply24vDrive1 := "i.A195AP1.A20QF3.PowerSupply24VDrive";
   //"ZUPS".tInputs.xDriveSupply1 := "i.A195AP1.A51QM1.DriveSupply";
   //"ZUPS".tInputs.xUPSEmLocMCC1201 := "i.A195AP1.A32SB1.EmergencyLocalizationUPS_MCC1201";
   //"ZUPS".tInputs.xUPSEmLocM203S_1 := "i.A401AP1.A32SB4.EmergencyLocalizationUPS_M203S";
   //"ZUPS".tInputs.xUPSEmLocM203S_2 := "i.A401AP1.A32SB5.EmergencyLocalizationUPS_M203S";

   "Z200".tInputs.xCPUAEnabled :="i.R150AP1.Selected CPU A";//"i.R195AP1.R125KA1 CPU A Enabled";
   "Z200".tInputs.xCPUBEnabled := "i.R150AP1.Selected CPU B";//"i.R195AP1.R125SA1Selection ON CPU B";
   "Z200".tInputs.xCPUARecognition := "i.R150AP1.Recognition CPU A";
   "Z200".tInputs.xCPUBRecognition := "i.R150AP1.Anomay Power supply  CPU B";
   "Z200".tInputs.xPowerSupply230vAux := "i.R195AP1.R11QF2/3.PowerFailure230VAuxiliary";
   "Z200".tInputs.xPowerSupply24vProt1 := "i.R195AP1.R18QF1.PowerFailure24VSuplly1";
   "Z200".tInputs.xPowerSupply24vProt2 := "i.R195AP1.R18QF2.PowerFailure24VSuplly2";
   "Z200".tInputs.xProtectionCommandsAnomalies := "i.R195AP1.R18QF3.PowerFailure24V_Commands";
   "Z200".tInputs.xProtectionCommandsInternalInput := "i.R195AP1.R18QF4.PowerFailure24V_Input";
   "Z200".tInputs.xFeedbackSwitch := "i.R195AP1.R125KA1CPU_A_Enabled";
   "Z200".tInputs.xFeedbackAbilitationCPU_B:="i.R195AP1.R125SA1SelectionOnCPU_B";
   "Z200".tInputs.xProtectionCommandsInternalOutput := "i.R195AP1.R18QF7.PowerSupply24VLogic";
   "Z200".tInputs.xProtectionCommandsExternalInput := "i.R195AP1.R18QF8.PowerSupply24VLogic";
   "Z200".tInputs.xRedundancy24vOk1 := "i.R195AP1.R18AP1.Redundacy24VOk";




   "Z200".tInputs.xCompressedAirPresence := "i.R195AP1.R427SSP1.CompressedAirPresenceCuttingBridge";



   "FB_Digitizer_1_V1_00_IDB".INPUTS.dEncCounter_count := "i_HSCInput_Count2".countValue;
   "FB_Digitizer_1_V1_00_IDB".INPUTS.xGlassPresence := "i.R195AP1.M216B1.GlassPresenceOnEncoder#1M216";

   "FB_Digitizer_2_V1_00_IDB".INPUTS.dEncCounter_count := "i_HSCInput_Count3".countValue;;
   "FB_Digitizer_2_V1_00_IDB".INPUTS.xGlassPresence := "i.R195AP1.M216B2.GlassPresenceOnEncoder#2M216";

   "FB_Oil_V1_00_IDB".INPUT.xPowerSupply := TRUE;
   "FB_Oil_V1_00_IDB".INPUT.xOilMaxLevel := "i.R195AP1.R427SL2.MaximumLevelOilTank";
   "FB_Oil_V1_00_IDB".INPUT.xOilMinLevel := "i.R195AP1.R427SL1.MinimumLevelOilTank";


   "FB_YCuts1_V1_00_IDB".IN_tIDeviceData := "i.MCC1256B1_IDevice";
   "FB_YCuts2_V1_00_IDB".IN_tIDeviceData := "i.MCC1256B2_IDevice";

   "FB_Markers_V1.00_IDB".IN_tIDeviceData := "i.MCC1204_IDeviceFromMarkers";

   "FB_BD_BreakPH_V1_00_IDB".INPUT.xPowerSupplyControl := TRUE;
   "FB_BD_BreakPH_V1_00_IDB".INPUT.xConnectorONOp := TRUE;
   "FB_BD_BreakPH_V1_00_IDB".INPUT.xConnectorONOppoOp := TRUE;


   "FB_BD_DigitizerPH_V1_00_IDB".INPUT.xPowerSupplyControl := TRUE;
   "FB_BD_DigitizerPH_V1_00_IDB".INPUT.xConnectorONOp := TRUE;
   "FB_BD_DigitizerPH_V1_00_IDB".INPUT.xConnectorONOppoOp := TRUE;

   "FB_BD_DigitizerPH_V1_00_IDB".INPUT.rgxPhotoStatus[0] := "i.R195AP1.M216B1.GlassPresenceOnEncoder#1M216";
   "FB_BD_DigitizerPH_V1_00_IDB".INPUT.rgxPhotoStatus[1] := "i.R195AP1.M216B2.GlassPresenceOnEncoder#2M216";
   "FB_BD_DigitizerPH_V1_00_IDB".INPUT.xButtonAlarmOFF:="FB_CommunicationZ300_V1.00_DB".IN_tIDeviceDataIN.Z200.IN_MCC1301."xE.E108.6";


   "FB_ManInsp_V1_00_IDB".INPUT.xPowerSupplyControl := TRUE;
   "FB_ManInsp_V1_00_IDB".INPUT.rgxQualityButtons[0] := "i.R195AP1.M212SB3.QualityB1";


   "FB_ManInsp_V1_00_IDB".INPUT.rgxDefectButtons[0] := "i.R195AP1.M212SB4.DefectButtonClass3";
   "FB_ManInsp_V1_00_IDB".INPUT.rgxDefectButtons[1] := "i.R195AP1.M212SB5.DefectButtonClass4";
   "FB_ManInsp_V1_00_IDB".INPUT.rgxDefectButtons[2] := "i.R195AP1.M212SB1.DefectButtonClass3";
   "FB_ManInsp_V1_00_IDB".INPUT.rgxDefectButtons[3] := "i.R195AP1.M212SB2.DefectButtonClass4";
   //"FB_ManInsp_V1_00_IDB".INPUT.rgxDefectButtons[2] := "i.A431AP1.A434SB4.M232.DefectButtonClass3_2";
   //"FB_ManInsp_V1_00_IDB".INPUT.rgxDefectButtons[3] := "i.A431AP1.A434SB4.M232.DefectButtonClass4_2";
   //"FB_ManInsp_V1_00_IDB".INPUT.rgxDefectButtons[4] := "i.R195AP1.M212SB1.DefectButtonClass3";
   //"FB_ManInsp_V1_00_IDB".INPUT.rgxDefectButtons[5] := "i.R195AP1.M212SB2.DefectButtonClass4";
   //"FB_ManInsp_V1_00_IDB".INPUT.rgxDefectButtons[6] := "i.A431AP1.A434SB7.M232.DefectButtonClass3_4";
   //"FB_ManInsp_V1_00_IDB".INPUT.rgxDefectButtons[7] := "i.A431AP1.A435SB1.M232.DefectButtonClass4_4";

   "FB_ISRA5D_IDB".IN_xScannerON := "i.R195AP1.SCANNER.ScannerOn";
   #TMP_xToAssign := "i.R195AP1.SCANNER.Scanner(1)";
END_REGION
END_FUNCTION

FUNCTION "InputTaskMedium" : Void   // FC10, LAD
{ S7_Optimized_Access := 'TRUE' }
VERSION : 0.1
BEGIN
END_FUNCTION

FUNCTION "InputZ201_Idevice" : Void   // FC30, LAD
{ S7_Optimized_Access := 'TRUE' }
VERSION : 0.1
   VAR_TEMP
      TMP_xToAssign : Bool;
   END_VAR
BEGIN

REGION Network 1 (SCL)
   "ZUPS".tInputs.xEmergencyONAreaUPS := "FB_CommunicationZ300_V1.00_DB".IN_tIDeviceDataIN.Z200.IN_MCC1201."xA.E80.4";
   "ZUPS".tInputs.xPowerSupply24vDrive1 := "FB_CommunicationZ300_V1.00_DB".IN_tIDeviceDataIN.Z200.IN_MCC1201."xA.E81.3";
   "ZUPS".tInputs.xDriveSupply1 := "FB_CommunicationZ300_V1.00_DB".IN_tIDeviceDataIN.Z200.IN_MCC1201."xA.E81.0";
   "ZUPS".tInputs.xUPSEmLocMCC1201 := "FB_CommunicationZ300_V1.00_DB".IN_tIDeviceDataIN.Z200.IN_MCC1201."xA.E80.6";
   "ZUPS".tInputs.xUPSEmLocM204S_1 := "FB_CommunicationZ300_V1.00_DB".IN_tIDeviceDataIN.Z200.IN_MCC1201."xA.E34.3";
   "ZUPS".tInputs.xUPSEmLocM204S_2 := "FB_CommunicationZ300_V1.00_DB".IN_tIDeviceDataIN.Z200.IN_MCC1201."xA.E35.1";

   "ZUPS".tInputs.xUPSEmLocCS4201 := "FB_CommunicationZ300_V1.00_DB".IN_tIDeviceDataIN.Z200.IN_MCC1201."xA.E38.0";



   "Z201".tInputs.xCPUAEnabled := "FB_CommunicationZ300_V1.00_DB".IN_tIDeviceDataIN.Z200.IN_MCC1201."xA.E20.0";
   "Z201".tInputs.xCPUBEnabled := "FB_CommunicationZ300_V1.00_DB".IN_tIDeviceDataIN.Z200.IN_MCC1201."xA.E20.1";
   "Z201".tInputs.xCPUARecognition := "FB_CommunicationZ300_V1.00_DB".IN_tIDeviceDataIN.Z200.IN_MCC1201."xA.E20.2";
   "Z201".tInputs.xCPUBRecognition :=  "FB_CommunicationZ300_V1.00_DB".IN_tIDeviceDataIN.Z200.IN_MCC1201."xA.E20.3";
   //"Z201".tInputs.xPowerSupply230vAux := "i.A195AP1.A10QF1/2.PowerFailure230VAuxiliary";
   "Z201".tInputs.xPowerSupply24vLogic1 := "FB_CommunicationZ300_V1.00_DB".IN_tIDeviceDataIN.Z200.IN_MCC1201."xA.E80.0";
   "Z201".tInputs.xPowerSupply24vLogic2 := "FB_CommunicationZ300_V1.00_DB".IN_tIDeviceDataIN.Z200.IN_MCC1201."xA.E80.1";
   "Z201".tInputs.xPowerSupply24vLogic3 := "FB_CommunicationZ300_V1.00_DB".IN_tIDeviceDataIN.Z200.IN_MCC1201."xA.E80.2";
   "Z201".tInputs.xPowerSupply24vLogic4 := "FB_CommunicationZ300_V1.00_DB".IN_tIDeviceDataIN.Z200.IN_MCC1201."xA.E80.3";
   "Z201".tInputs.xPowerSuppluyOut24vUnderUpsEmOk := "FB_CommunicationZ300_V1.00_DB".IN_tIDeviceDataIN.Z200.IN_MCC1201."xA.E80.2"AND"FB_CommunicationZ300_V1.00_DB".IN_tIDeviceDataIN.Z200.IN_MCC1201."xA.E80.4"AND "CU_A250AP1_IDB".STC_tPZD_CU.tR.tE_DIGITAL.x8 ;
   "Z201".tInputs.xPowerSuppluyOut24vUnderEmOk := "FB_CommunicationZ300_V1.00_DB".IN_tIDeviceDataIN.Z200.IN_MCC1201."xA.E80.5"AND "FB_CommunicationZ300_V1.00_DB".IN_tIDeviceDataIN.Z200.IN_MCC1201."xA.E80.3"AND"CU_A260AP1_IDB".STC_tPZD_CU.tR.tE_DIGITAL.x8 ;
   "Z201".tInputs.xMainEmergencyON := "FB_CommunicationZ300_V1.00_DB".IN_tIDeviceDataIN.Z200.IN_MCC1201."xA.E80.5";
   "Z201".tInputs.xM216FanFeedback := "FB_CommunicationZ300_V1.00_DB".IN_tIDeviceDataIN.Z200.IN_MCC1201."xA.E81.7";
   "Z201".tInputs.xM216FanProtection := "FB_CommunicationZ300_V1.00_DB".IN_tIDeviceDataIN.Z200.IN_MCC1201."xA.E81.6";

   "Z201".tInputs.xPowerSupply24vDrive2 := "FB_CommunicationZ300_V1.00_DB".IN_tIDeviceDataIN.Z200.IN_MCC1201."xA.E81.4";
   "Z201".tInputs.xEmLocMCC1201 := "FB_CommunicationZ300_V1.00_DB".IN_tIDeviceDataIN.Z200.IN_MCC1201."xA.E80.6";
   "Z201".tInputs.xEmergencyONArea201 :=  "FB_CommunicationZ300_V1.00_DB".IN_tIDeviceDataIN.Z200.IN_MCC1201."xA.E33.7"OR"FB_CommunicationZ300_V1.00_DB".IN_tIDeviceDataIN.Z200.IN_MCC1201."xA.E34.4"OR"FB_CommunicationZ300_V1.00_DB".IN_tIDeviceDataIN.Z200.IN_MCC1201."xA.E36.4"OR"FB_CommunicationZ300_V1.00_DB".IN_tIDeviceDataIN.Z200.IN_MCC1201."xA.E36.5"OR"FB_CommunicationZ300_V1.00_DB".IN_tIDeviceDataIN.Z200.IN_MCC1201."xA.E37.0"OR"FB_CommunicationZ300_V1.00_DB".IN_tIDeviceDataIN.Z200.IN_MCC1201."xA.E37.1"OR"FB_CommunicationZ300_V1.00_DB".IN_tIDeviceDataIN.Z200.IN_MCC1201."xA.E37.4"OR"FB_CommunicationZ300_V1.00_DB".IN_tIDeviceDataIN.Z200.IN_MCC1201."xA.E37.5"OR"FB_CommunicationZ300_V1.00_DB".IN_tIDeviceDataIN.Z200.IN_MCC1201."xA.E38.1"OR"FB_CommunicationZ300_V1.00_DB".IN_tIDeviceDataIN.Z200.IN_MCC1201."xA.E80.6";

   "Z201".tInputs.xSBchipBlowerON_M209:="FB_CommunicationZ300_V1.00_DB".IN_tIDeviceDataIN.Z200.IN_MCC1201."xA.E36.2";

   //"Z201".tInputs.xEmergencyONArea301 := "i.MCC1301.E406AP1.M302SB1.EmergencyLocalization" OR "i.MCC1301.E406AP1.M302SB2.EmergencyLocalization" OR"i.MCC1301.E406AP1.M306SB1.EmergencyLocalization" OR"i.MCC1301.E406AP1.M312SSB1.EmergencyLocalization" OR"i.MCC1301.E406AP1.M312SSB2.EmergencyLocalization"OR "i.MCC1301.E405AP1.E121SB1.EmergencyLocalization" ;
   //"Z201".tInputs.xEmergencyONArea302 := "i.MCC1302.F405AP1.M317SSB1.EmergencyLocalization"OR "i.MCC1302.F405AP1.M317SSB2.EmergencyLocalization" OR"i.MCC1302.F405AP1.M319SB1.EmergencyLocalization" OR"i.MCC1302.F405AP1.M320SSB1.EmergencyLocalization" OR"i.MCC1302.F405AP1.M320SSB2.EmergencyLocalization" OR"i.MCC1302.F405AP1.M325SSB1.EmergencyLocalization"OR "i.MCC1302.F405AP1.M325SSB2.EmergencyLocalization"OR "i.MCC1302.F405AP1.F121SB1.EmergencyLocalization";
   //"Z201".tInputs.xEmergencyONArea303 := "i.MCC1303.G195AP1.G32SB1.EmergencyLocalization"OR "i.MCC1303.G195AP1.M323SB1.EmergencyLocalization" OR"i.MCC1303.G195AP1.M323SB2.EmergencyLocalization" ;
   //"Z201".tInputs.xEmergencyONArea601 := "i.A195AP1.A38KE2.EmergencyArea601ON";
   //"Z201".tInputs.xEmergencyONArea701 := "i.A195AP1.A39KE1.EmergencyArea701ON";
   "Z201".tInputs.xDriveSupply2 := "FB_CommunicationZ300_V1.00_DB".IN_tIDeviceDataIN.Z200.IN_MCC1201."xA.E81.1";
   "Z201".tInputs.xSBResetAnomalyZ200 := "FB_CommunicationZ300_V1.00_DB".IN_tIDeviceDataIN.Z200.IN_MCC1301."xE.E108.0";
   "Z201".tInputs.xEmLocCS4201 := "FB_CommunicationZ300_V1.00_DB".IN_tIDeviceDataIN.Z200.IN_MCC1201."xA.E38.4";
   "Z201".tInputs.xEmLocM204S_1 := "FB_CommunicationZ300_V1.00_DB".IN_tIDeviceDataIN.Z200.IN_MCC1201."xA.E34.4";
   "Z201".tInputs.xEmLocM204S_2 := "FB_CommunicationZ300_V1.00_DB".IN_tIDeviceDataIN.Z200.IN_MCC1201."xA.E35.2";
   "Z201".tInputs.xEmLocM211_1 := "FB_CommunicationZ300_V1.00_DB".IN_tIDeviceDataIN.Z200.IN_MCC1201."xA.E36.4";
   "Z201".tInputs.xEmLocM211_2 :=  "FB_CommunicationZ300_V1.00_DB".IN_tIDeviceDataIN.Z200.IN_MCC1201."xA.E36.5";
   "Z201".tInputs.xEmLocM214_1 := "FB_CommunicationZ300_V1.00_DB".IN_tIDeviceDataIN.Z200.IN_MCC1201."xA.E37.0";
   "Z201".tInputs.xEmLocM214_2 := "FB_CommunicationZ300_V1.00_DB".IN_tIDeviceDataIN.Z200.IN_MCC1201."xA.E37.1";
   "Z201".tInputs.xEmLocM218_1 := "FB_CommunicationZ300_V1.00_DB".IN_tIDeviceDataIN.Z200.IN_MCC1201."xA.E37.4";
   "Z201".tInputs.xEmLocM218_2:= "FB_CommunicationZ300_V1.00_DB".IN_tIDeviceDataIN.Z200.IN_MCC1201."xA.E37.5";
   "Z201".tInputs.xEmLocCS4202 := "FB_CommunicationZ300_V1.00_DB".IN_tIDeviceDataIN.Z200.IN_MCC1201."xA.E38.1";